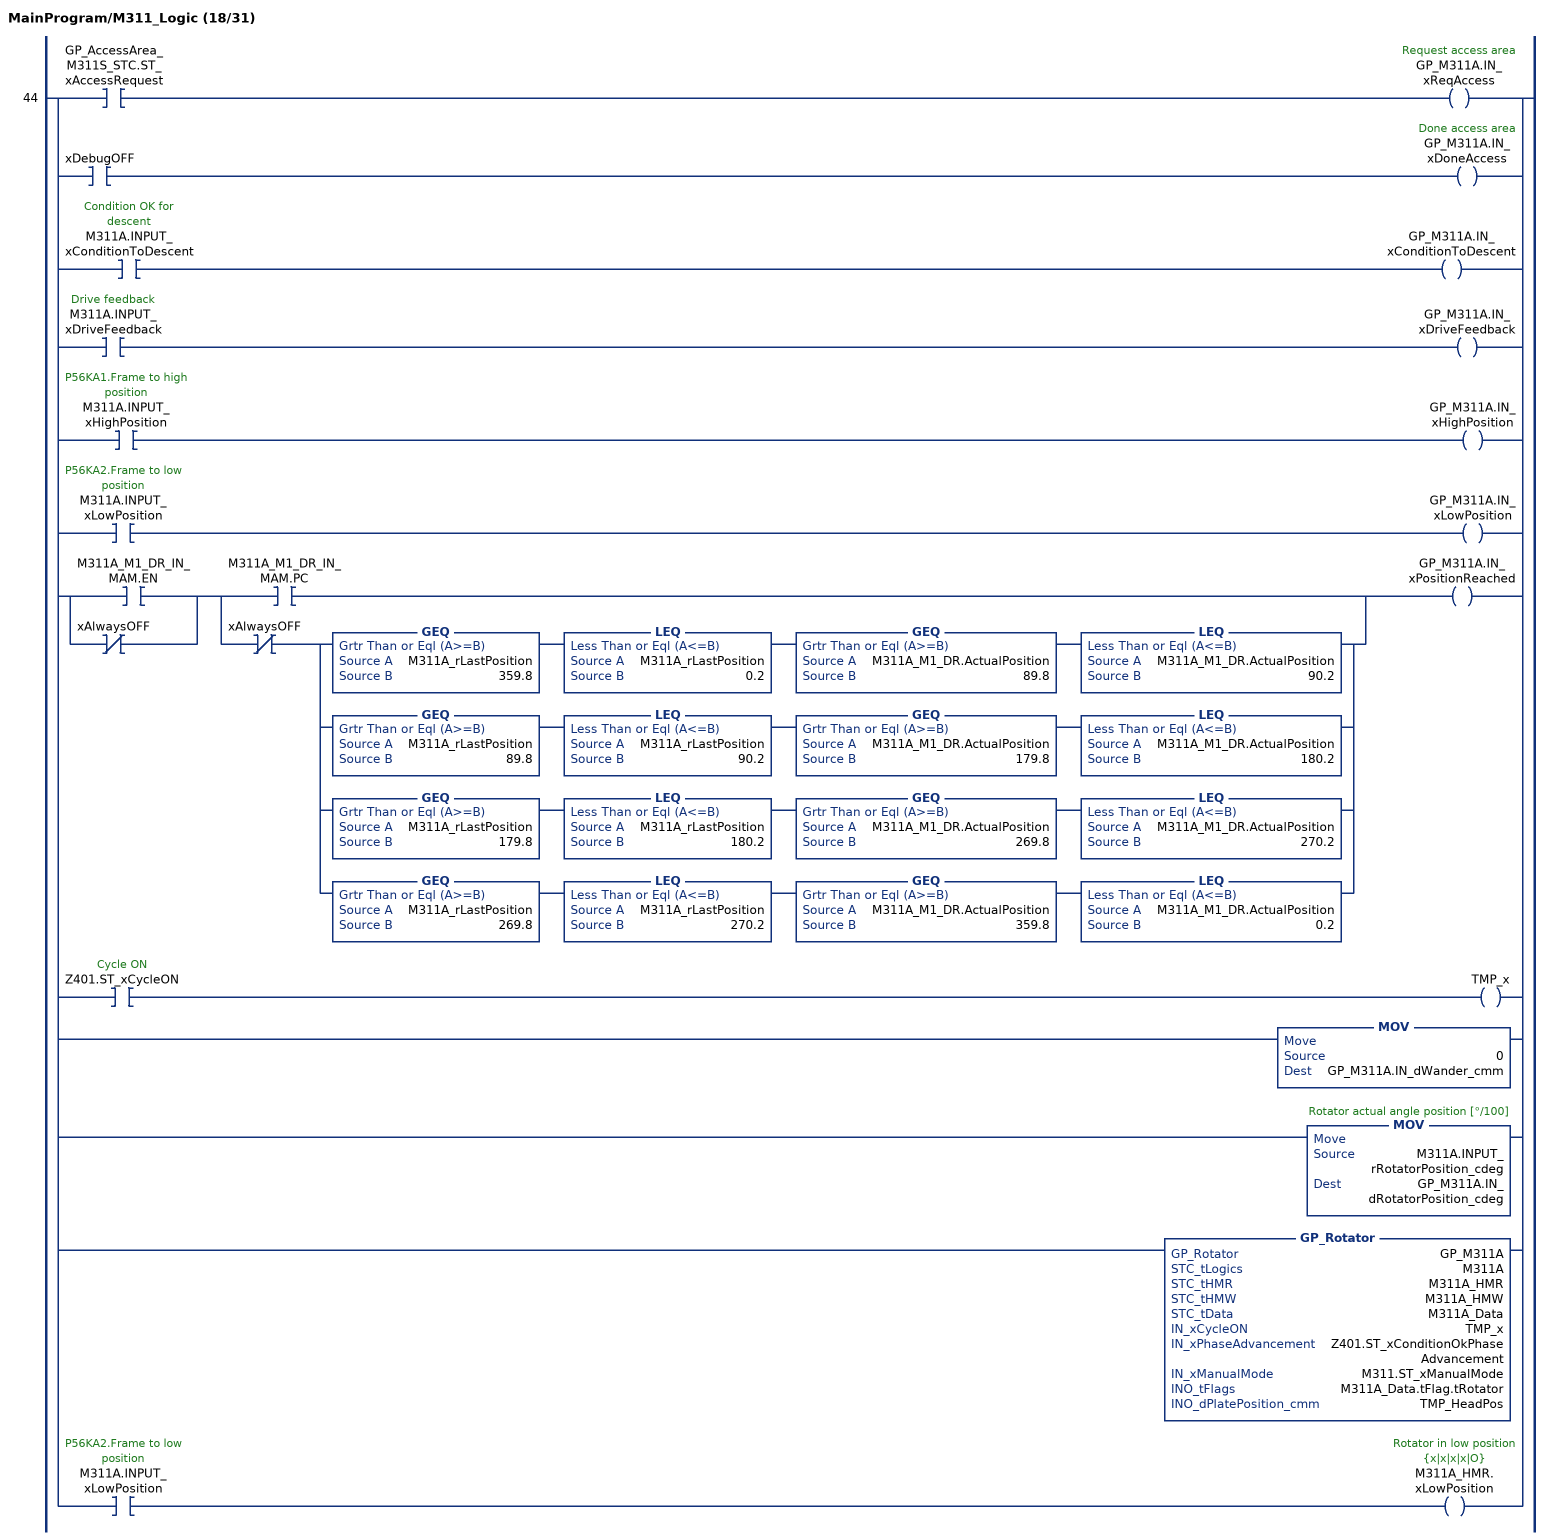
   44: [XIC(GP_AccessArea_M311S_STC.ST_xAccessRequest) OTE(GP_M311A.IN_xReqAccess) ,XIC(xDebugOFF) OTE(GP_M311A.IN_xDoneAccess) ,XIC(M311A.INPUT_xConditionToDescent) OTE(GP_M311A.IN_xConditionToDescent) ,XIC(M311A.INPUT_xDriveFeedback) OTE(GP_M311A.IN_xDriveFeedback) ,XIC(M311A.INPUT_xHighPosition) OTE(GP_M311A.IN_xHighPosition) ,XIC(M311A.INPUT_xLowPosition) OTE(GP_M311A.IN_xLowPosition) ,[XIC(M311A_M1_DR_IN_MAM.EN) ,XIO(xAlwaysOFF) ] [XIC(M311A_M1_DR_IN_MAM.PC) ,XIO(xAlwaysOFF) [GEQ(M311A_rLastPosition,359.8) LEQ(M311A_rLastPosition,0.2) GEQ(M311A_M1_DR.ActualPosition,89.8) LEQ(M311A_M1_DR.ActualPosition,90.2) ,GEQ(M311A_rLastPosition,89.8) LEQ(M311A_rLastPosition,90.2) GEQ(M311A_M1_DR.ActualPosition,179.8) LEQ(M311A_M1_DR.ActualPosition,180.2) ,GEQ(M311A_rLastPosition,179.8) LEQ(M311A_rLastPosition,180.2) GEQ(M311A_M1_DR.ActualPosition,269.8) LEQ(M311A_M1_DR.ActualPosition,270.2) ,GEQ(M311A_rLastPosition,269.8) LEQ(M311A_rLastPosition,270.2) GEQ(M311A_M1_DR.ActualPosition,359.8) LEQ(M311A_M1_DR.ActualPosition,0.2) ] ] OTE(GP_M311A.IN_xPositionReached) ,XIC(Z401.ST_xCycleON) OTE(TMP_x) ,MOV(0,GP_M311A.IN_dWander_cmm) ,MOV(M311A.INPUT_rRotatorPosition_cdeg,GP_M311A.IN_dRotatorPosition_cdeg) ,GP_Rotator(GP_M311A,M311A,M311A_HMR,M311A_HMW,M311A_Data,TMP_x,Z401.ST_xConditionOkPhaseAdvancement,M311.ST_xManualMode,M311A_Data.tFlag.tRotator,TMP_HeadPos) ,XIC(M311A.INPUT_xLowPosition) OTE(M311A_HMR.xLowPosition) ];
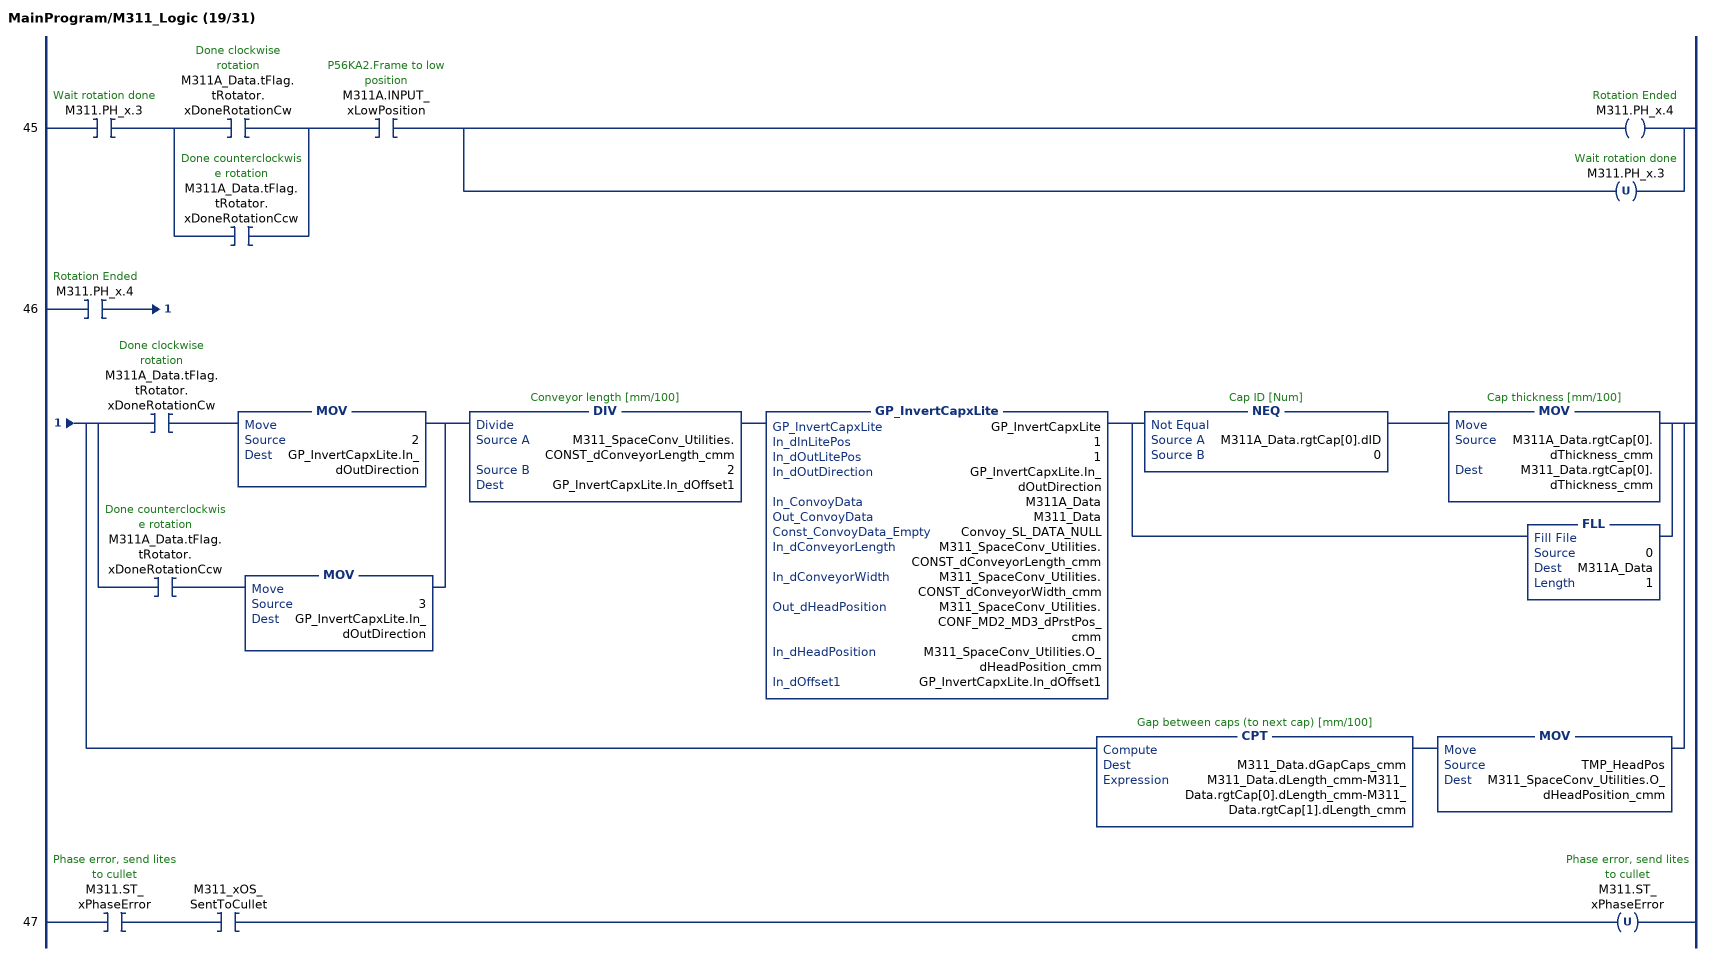
   45: XIC(M311.PH_x.3)[XIC(M311A_Data.tFlag.tRotator.xDoneRotationCw) ,XIC(M311A_Data.tFlag.tRotator.xDoneRotationCcw) ]XIC(M311A.INPUT_xLowPosition)[OTE(M311.PH_x.4) ,OTU(M311.PH_x.3) ];
   46: XIC(M311.PH_x.4)[[XIC(M311A_Data.tFlag.tRotator.xDoneRotationCw) MOV(2,GP_InvertCapxLite.In_dOutDirection) ,XIC(M311A_Data.tFlag.tRotator.xDoneRotationCcw) MOV(3,GP_InvertCapxLite.In_dOutDirection) ] DIV(M311_SpaceConv_Utilities.CONST_dConveyorLength_cmm,2,GP_InvertCapxLite.In_dOffset1) GP_InvertCapxLite(GP_InvertCapxLite,1,1,GP_InvertCapxLite.In_dOutDirection,M311A_Data,M311_Data,Convoy_SL_DATA_NULL,M311_SpaceConv_Utilities.CONST_dConveyorLength_cmm,M311_SpaceConv_Utilities.CONST_dConveyorWidth_cmm,M311_SpaceConv_Utilities.CONF_MD2_MD3_dPrstPos_cmm,M311_SpaceConv_Utilities.O_dHeadPosition_cmm,GP_InvertCapxLite.In_dOffset1) [NEQ(M311A_Data.rgtCap[0].dID,0) MOV(M311A_Data.rgtCap[0].dThickness_cmm,M311_Data.rgtCap[0].dThickness_cmm) ,FLL(0,M311A_Data,1) ] ,CPT(M311_Data.dGapCaps_cmm,M311_Data.dLength_cmm-M311_Data.rgtCap[0].dLength_cmm-M311_Data.rgtCap[1].dLength_cmm) MOV(TMP_HeadPos,M311_SpaceConv_Utilities.O_dHeadPosition_cmm) ];
   47: XIC(M311.ST_xPhaseError)XIC(M311_xOS_SentToCullet)OTU(M311.ST_xPhaseError);
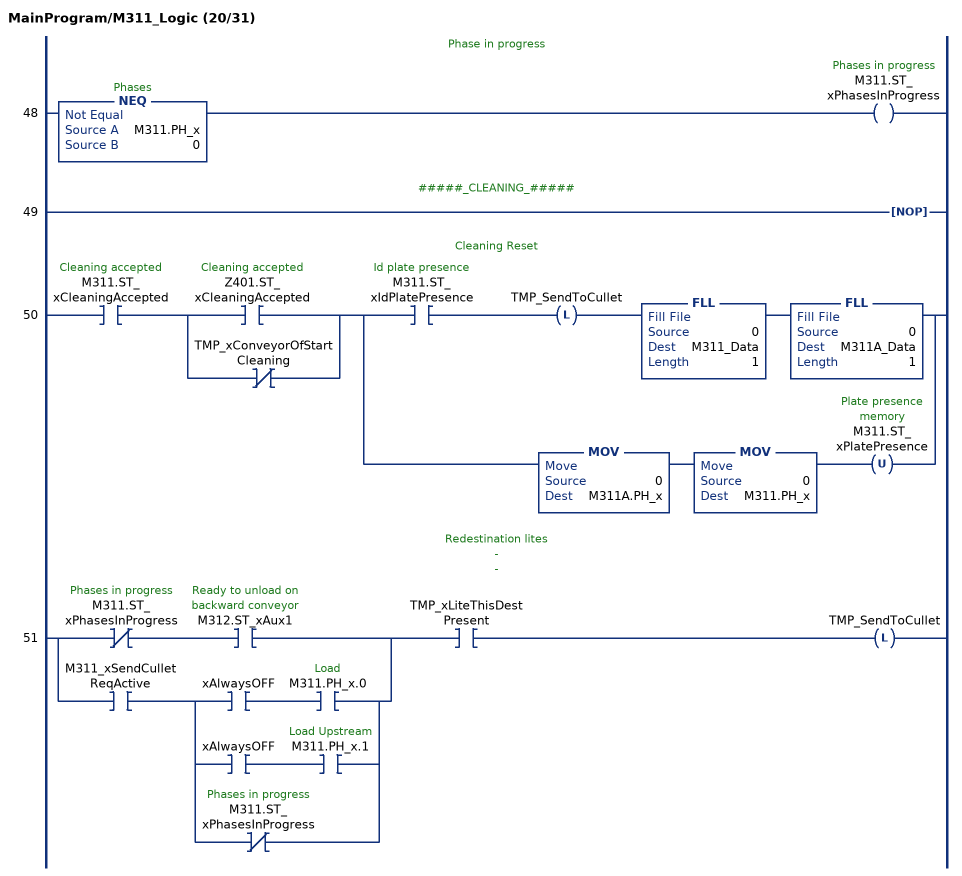
   // Phase in progress
   48: NEQ(M311.PH_x,0)OTE(M311.ST_xPhasesInProgress);
   // #####_CLEANING_#####
   49: NOP();
   // Cleaning Reset
   50: XIC(M311.ST_xCleaningAccepted)[XIC(Z401.ST_xCleaningAccepted) ,XIO(TMP_xConveyorOfStartCleaning) ][XIC(M311.ST_xIdPlatePresence) OTL(TMP_SendToCullet) FLL(0,M311_Data,1) FLL(0,M311A_Data,1) ,MOV(0,M311A.PH_x) MOV(0,M311.PH_x) OTU(M311.ST_xPlatePresence) ];
   // Redestination lites
   // -
   // -
   51: [XIO(M311.ST_xPhasesInProgress) XIC(M312.ST_xAux1) ,XIC(M311_xSendCulletReqActive) [XIC(xAlwaysOFF) XIC(M311.PH_x.0) ,XIC(xAlwaysOFF) XIC(M311.PH_x.1) ,XIO(M311.ST_xPhasesInProgress) ] ]XIC(TMP_xLiteThisDestPresent)OTL(TMP_SendToCullet);
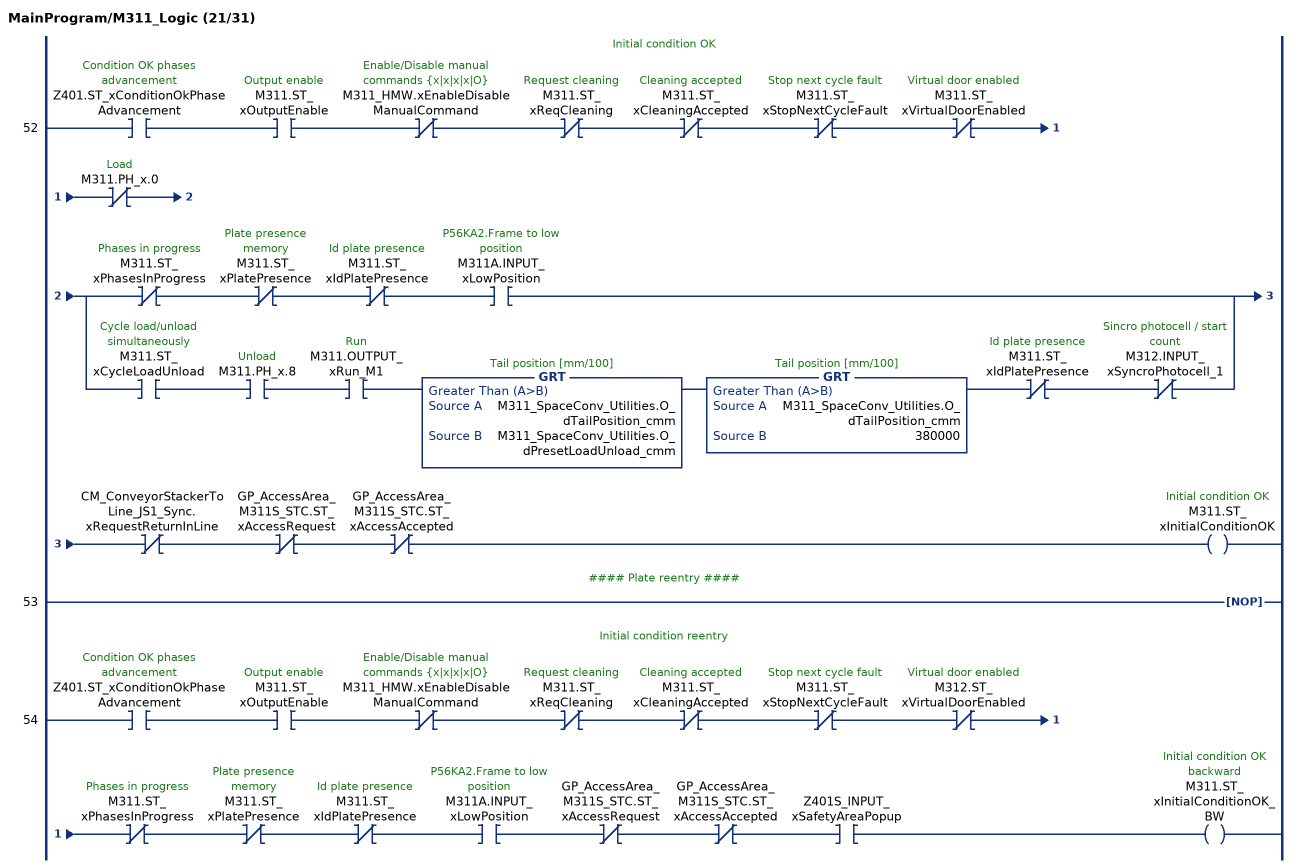
   // Initial condition OK
   52: XIC(Z401.ST_xConditionOkPhaseAdvancement)XIC(M311.ST_xOutputEnable)XIO(M311_HMW.xEnableDisableManualCommand)XIO(M311.ST_xReqCleaning)XIO(M311.ST_xCleaningAccepted)XIO(M311.ST_xStopNextCycleFault)XIO(M311.ST_xVirtualDoorEnabled)XIO(M311.PH_x.0)[XIO(M311.ST_xPhasesInProgress) XIO(M311.ST_xPlatePresence) XIO(M311.ST_xIdPlatePresence) XIC(M311A.INPUT_xLowPosition) ,XIC(M311.ST_xCycleLoadUnload) XIC(M311.PH_x.8) XIC(M311.OUTPUT_xRun_M1) GRT(M311_SpaceConv_Utilities.O_dTailPosition_cmm,M311_SpaceConv_Utilities.O_dPresetLoadUnload_cmm) GRT(M311_SpaceConv_Utilities.O_dTailPosition_cmm,380000) XIO(M311.ST_xIdPlatePresence) XIO(M312.INPUT_xSyncroPhotocell_1) ]XIO(CM_ConveyorStackerToLine_JS1_Sync.xRequestReturnInLine)XIO(GP_AccessArea_M311S_STC.ST_xAccessRequest)XIO(GP_AccessArea_M311S_STC.ST_xAccessAccepted)OTE(M311.ST_xInitialConditionOK);
   // #### Plate reentry ####
   53: NOP();
   // Initial condition reentry
   54: XIC(Z401.ST_xConditionOkPhaseAdvancement)XIC(M311.ST_xOutputEnable)XIO(M311_HMW.xEnableDisableManualCommand)XIO(M311.ST_xReqCleaning)XIO(M311.ST_xCleaningAccepted)XIO(M311.ST_xStopNextCycleFault)XIO(M312.ST_xVirtualDoorEnabled)XIO(M311.ST_xPhasesInProgress)XIO(M311.ST_xPlatePresence)XIO(M311.ST_xIdPlatePresence)XIC(M311A.INPUT_xLowPosition)XIO(GP_AccessArea_M311S_STC.ST_xAccessRequest)XIO(GP_AccessArea_M311S_STC.ST_xAccessAccepted)XIC(Z401S_INPUT_xSafetyAreaPopup)OTE(M311.ST_xInitialConditionOK_BW);
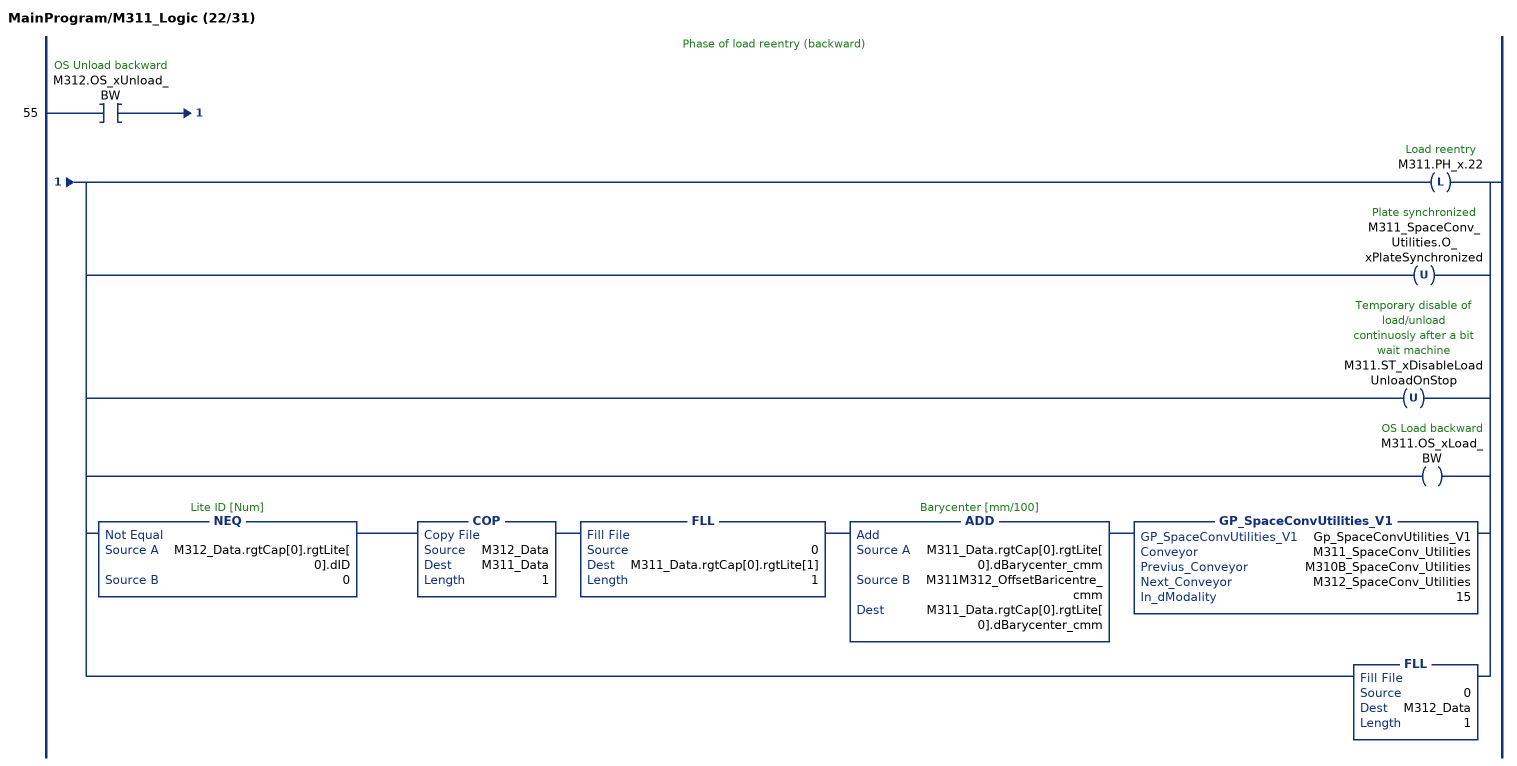
   // Phase of load reentry (backward)
   55: XIC(M312.OS_xUnload_BW)[OTL(M311.PH_x.22) ,OTU(M311_SpaceConv_Utilities.O_xPlateSynchronized) ,OTU(M311.ST_xDisableLoadUnloadOnStop) ,OTE(M311.OS_xLoad_BW) ,NEQ(M312_Data.rgtCap[0].rgtLite[0].dID,0) COP(M312_Data,M311_Data,1) FLL(0,M311_Data.rgtCap[0].rgtLite[1],1) ADD(M311_Data.rgtCap[0].rgtLite[0].dBarycenter_cmm,M311M312_OffsetBaricentre_cmm,M311_Data.rgtCap[0].rgtLite[0].dBarycenter_cmm) GP_SpaceConvUtilities_V1(Gp_SpaceConvUtilities_V1,M311_SpaceConv_Utilities,M310B_SpaceConv_Utilities,M312_SpaceConv_Utilities,15) ,FLL(0,M312_Data,1) ];
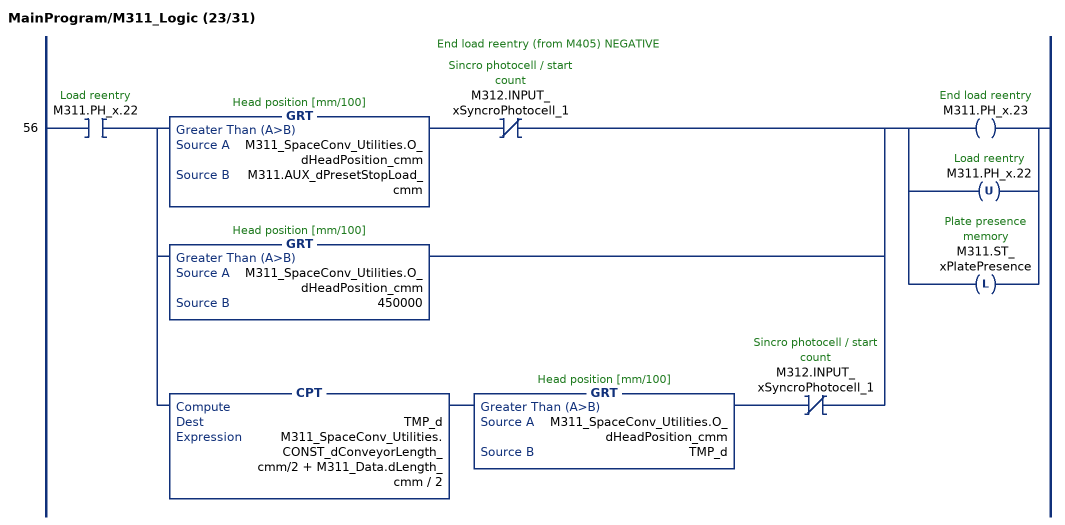
   // End load reentry (from M405) NEGATIVE
   56: XIC(M311.PH_x.22)[[GRT(M311_SpaceConv_Utilities.O_dHeadPosition_cmm,M311.AUX_dPresetStopLoad_cmm) XIO(M312.INPUT_xSyncroPhotocell_1) ,GRT(M311_SpaceConv_Utilities.O_dHeadPosition_cmm,450000) ] ,CPT(TMP_d,M311_SpaceConv_Utilities.CONST_dConveyorLength_cmm/2 + M311_Data.dLength_cmm / 2) GRT(M311_SpaceConv_Utilities.O_dHeadPosition_cmm,TMP_d) XIO(M312.INPUT_xSyncroPhotocell_1) ][OTE(M311.PH_x.23) ,OTU(M311.PH_x.22) ,OTL(M311.ST_xPlatePresence) ];
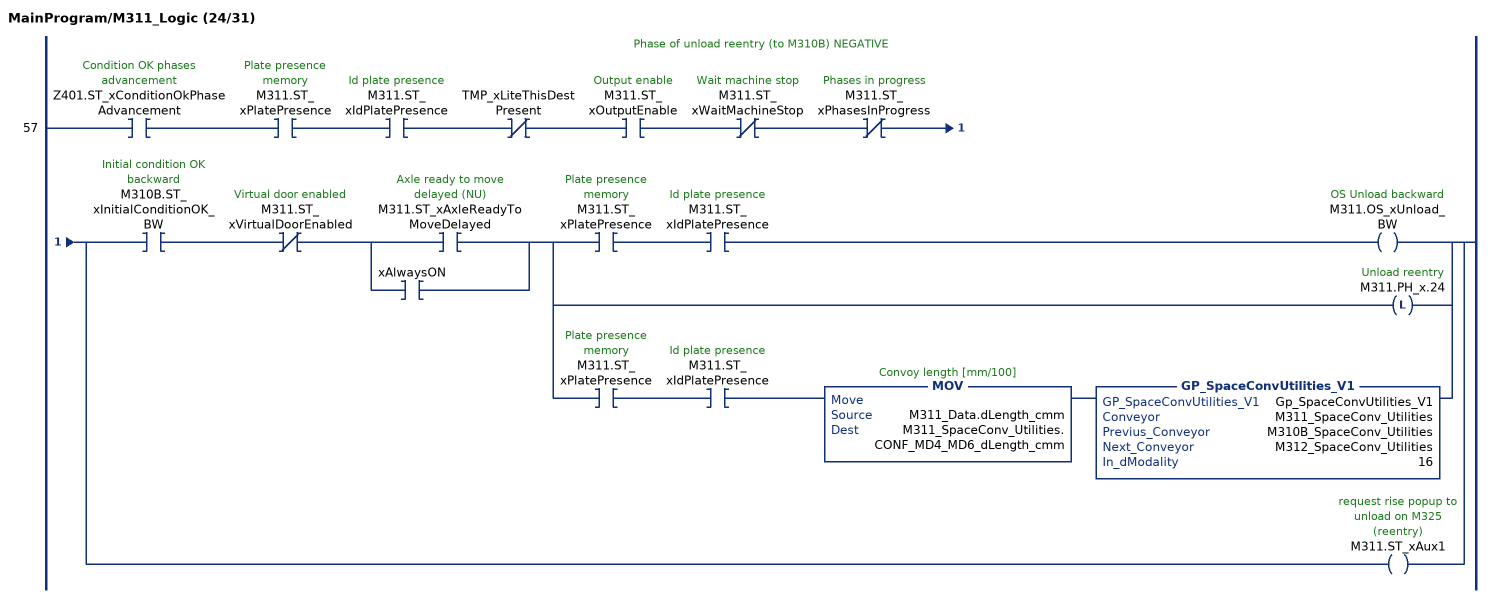
   // Phase of unload reentry (to M310B) NEGATIVE
   57: XIC(Z401.ST_xConditionOkPhaseAdvancement)XIC(M311.ST_xPlatePresence)XIC(M311.ST_xIdPlatePresence)XIO(TMP_xLiteThisDestPresent)XIC(M311.ST_xOutputEnable)XIO(M311.ST_xWaitMachineStop)XIO(M311.ST_xPhasesInProgress)[XIC(M310B.ST_xInitialConditionOK_BW) XIO(M311.ST_xVirtualDoorEnabled) [XIC(M311.ST_xAxleReadyToMoveDelayed) ,XIC(xAlwaysON) ] [XIC(M311.ST_xPlatePresence) XIC(M311.ST_xIdPlatePresence) OTE(M311.OS_xUnload_BW) ,OTL(M311.PH_x.24) ,XIC(M311.ST_xPlatePresence) XIC(M311.ST_xIdPlatePresence) MOV(M311_Data.dLength_cmm,M311_SpaceConv_Utilities.CONF_MD4_MD6_dLength_cmm) GP_SpaceConvUtilities_V1(Gp_SpaceConvUtilities_V1,M311_SpaceConv_Utilities,M310B_SpaceConv_Utilities,M312_SpaceConv_Utilities,16) ] ,OTE(M311.ST_xAux1) ];
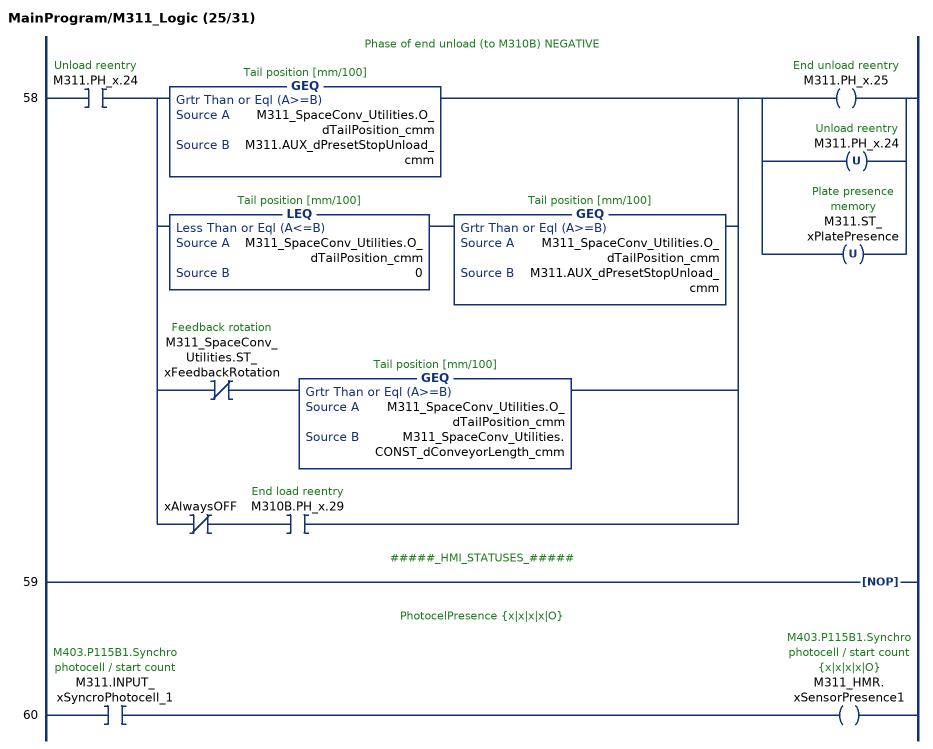
   // Phase of end unload (to M310B) NEGATIVE
   58: XIC(M311.PH_x.24)[[GEQ(M311_SpaceConv_Utilities.O_dTailPosition_cmm,M311.AUX_dPresetStopUnload_cmm) ,LEQ(M311_SpaceConv_Utilities.O_dTailPosition_cmm,0) GEQ(M311_SpaceConv_Utilities.O_dTailPosition_cmm,M311.AUX_dPresetStopUnload_cmm) ] ,XIO(M311_SpaceConv_Utilities.ST_xFeedbackRotation) GEQ(M311_SpaceConv_Utilities.O_dTailPosition_cmm,M311_SpaceConv_Utilities.CONST_dConveyorLength_cmm) ,XIO(xAlwaysOFF) XIC(M310B.PH_x.29) ][OTE(M311.PH_x.25) ,OTU(M311.PH_x.24) ,OTU(M311.ST_xPlatePresence) ];
   // #####_HMI_STATUSES_#####
   59: NOP();
   // PhotocelPresence {x|x|x|x|O}
   60: XIC(M311.INPUT_xSyncroPhotocell_1)OTE(M311_HMR.xSensorPresence1);
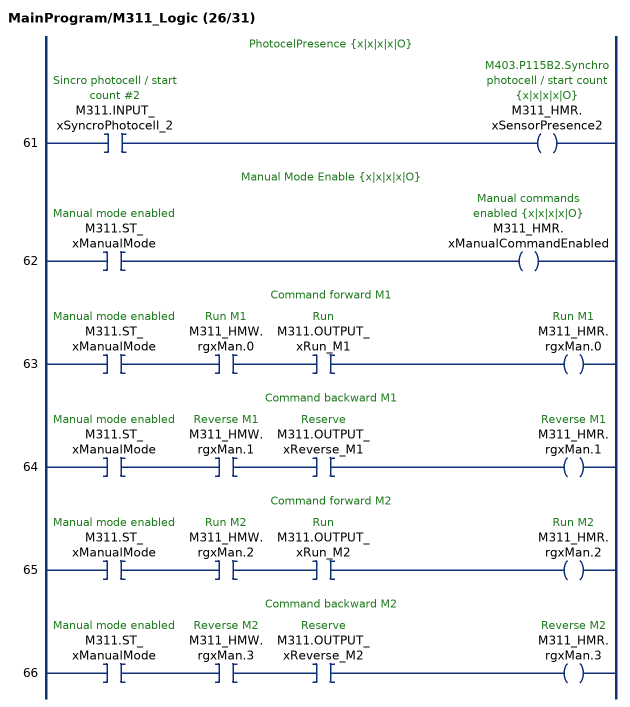
   // PhotocelPresence {x|x|x|x|O}
   61: XIC(M311.INPUT_xSyncroPhotocell_2)OTE(M311_HMR.xSensorPresence2);
   // Manual Mode Enable {x|x|x|x|O}
   62: XIC(M311.ST_xManualMode)OTE(M311_HMR.xManualCommandEnabled);
   // Command forward M1
   63: XIC(M311.ST_xManualMode)XIC(M311_HMW.rgxMan.0)XIC(M311.OUTPUT_xRun_M1)OTE(M311_HMR.rgxMan.0);
   // Command backward M1
   64: XIC(M311.ST_xManualMode)XIC(M311_HMW.rgxMan.1)XIC(M311.OUTPUT_xReverse_M1)OTE(M311_HMR.rgxMan.1);
   // Command forward M2
   65: XIC(M311.ST_xManualMode)XIC(M311_HMW.rgxMan.2)XIC(M311.OUTPUT_xRun_M2)OTE(M311_HMR.rgxMan.2);
   // Command backward M2
   66: XIC(M311.ST_xManualMode)XIC(M311_HMW.rgxMan.3)XIC(M311.OUTPUT_xReverse_M2)OTE(M311_HMR.rgxMan.3);
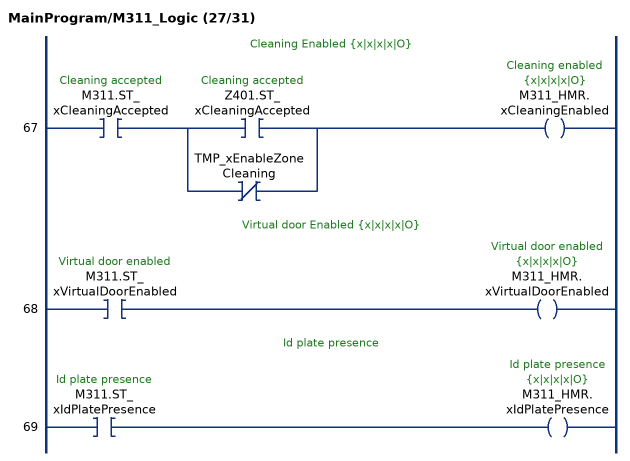
   // Cleaning Enabled {x|x|x|x|O}
   67: XIC(M311.ST_xCleaningAccepted)[XIC(Z401.ST_xCleaningAccepted) ,XIO(TMP_xEnableZoneCleaning) ]OTE(M311_HMR.xCleaningEnabled);
   // Virtual door Enabled {x|x|x|x|O}
   68: XIC(M311.ST_xVirtualDoorEnabled)OTE(M311_HMR.xVirtualDoorEnabled);
   // Id plate presence
   69: XIC(M311.ST_xIdPlatePresence)OTE(M311_HMR.xIdPlatePresence);
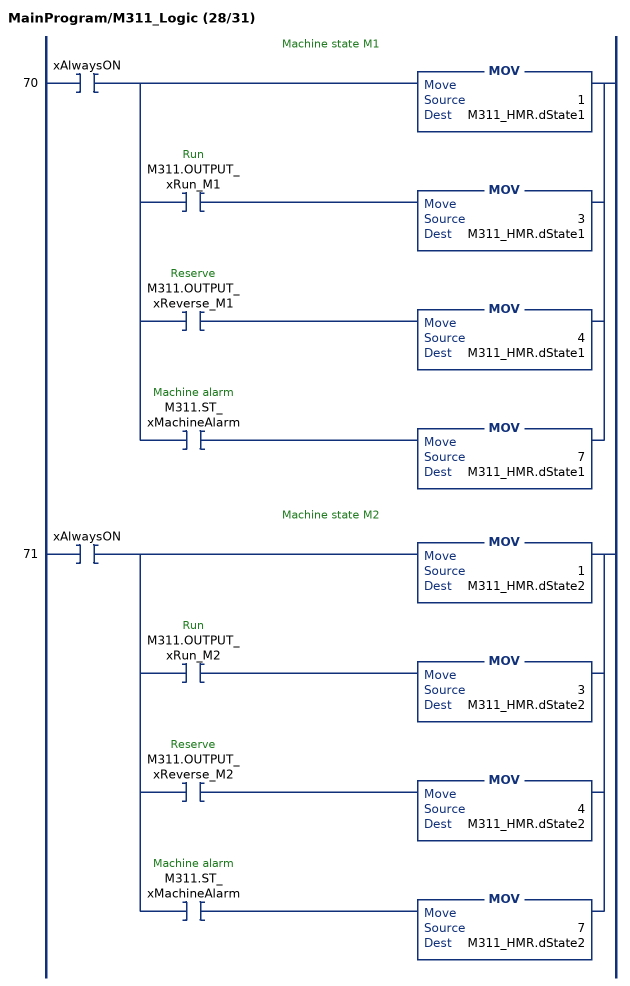
   // Machine state M1
   70: XIC(xAlwaysON)[MOV(1,M311_HMR.dState1) ,XIC(M311.OUTPUT_xRun_M1) MOV(3,M311_HMR.dState1) ,XIC(M311.OUTPUT_xReverse_M1) MOV(4,M311_HMR.dState1) ,XIC(M311.ST_xMachineAlarm) MOV(7,M311_HMR.dState1) ];
   // Machine state M2
   71: XIC(xAlwaysON)[MOV(1,M311_HMR.dState2) ,XIC(M311.OUTPUT_xRun_M2) MOV(3,M311_HMR.dState2) ,XIC(M311.OUTPUT_xReverse_M2) MOV(4,M311_HMR.dState2) ,XIC(M311.ST_xMachineAlarm) MOV(7,M311_HMR.dState2) ];
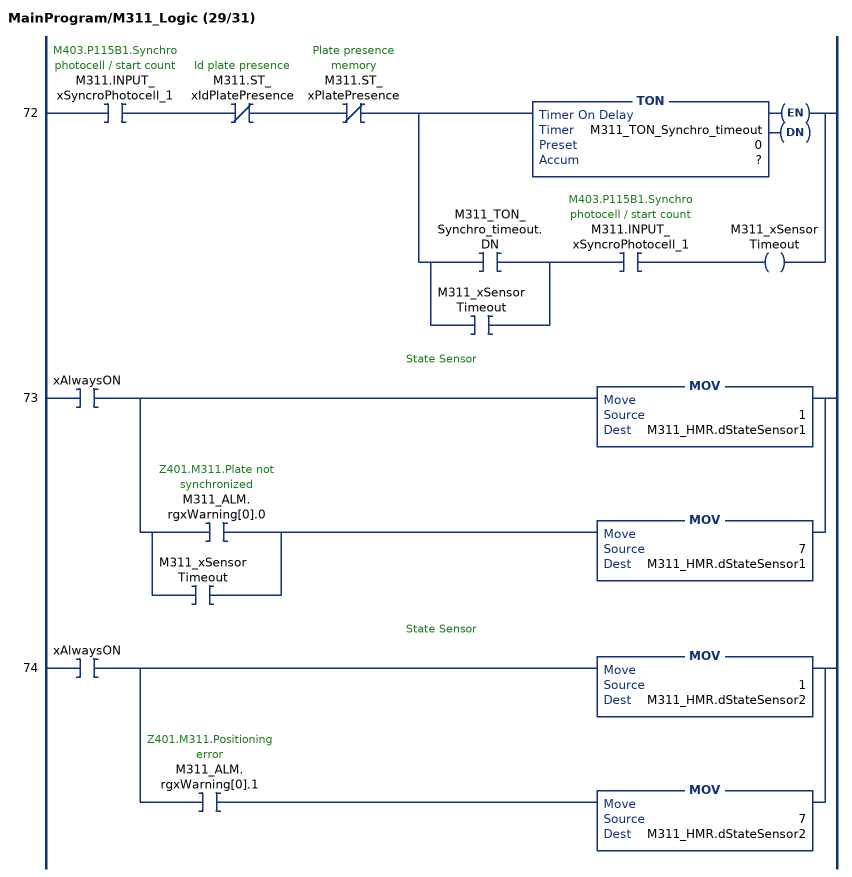
   72: XIC(M311.INPUT_xSyncroPhotocell_1)XIO(M311.ST_xIdPlatePresence)XIO(M311.ST_xPlatePresence)[TON(M311_TON_Synchro_timeout,?,?) ,[XIC(M311_TON_Synchro_timeout.DN) ,XIC(M311_xSensorTimeout) ] XIC(M311.INPUT_xSyncroPhotocell_1) OTE(M311_xSensorTimeout) ];
   // State Sensor
   73: XIC(xAlwaysON)[MOV(1,M311_HMR.dStateSensor1) ,[XIC(M311_ALM.rgxWarning[0].0) ,XIC(M311_xSensorTimeout) ] MOV(7,M311_HMR.dStateSensor1) ];
   // State Sensor
   74: XIC(xAlwaysON)[MOV(1,M311_HMR.dStateSensor2) ,XIC(M311_ALM.rgxWarning[0].1) MOV(7,M311_HMR.dStateSensor2) ];
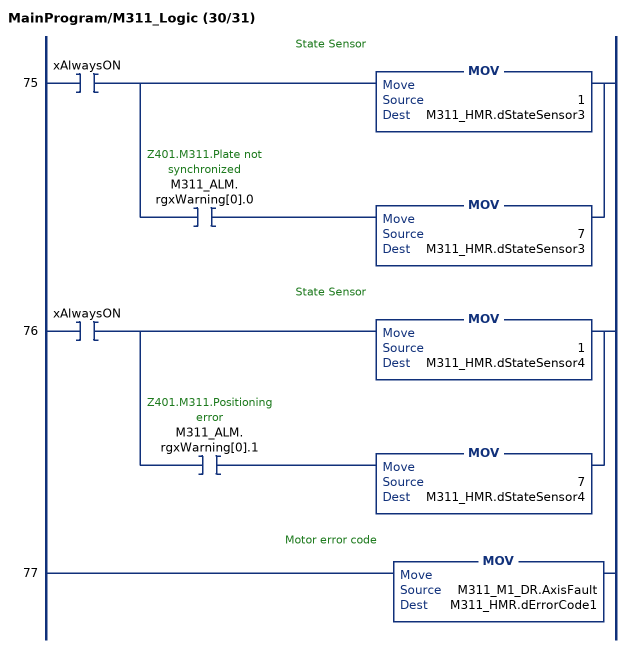
   // State Sensor
   75: XIC(xAlwaysON)[MOV(1,M311_HMR.dStateSensor3) ,XIC(M311_ALM.rgxWarning[0].0) MOV(7,M311_HMR.dStateSensor3) ];
   // State Sensor
   76: XIC(xAlwaysON)[MOV(1,M311_HMR.dStateSensor4) ,XIC(M311_ALM.rgxWarning[0].1) MOV(7,M311_HMR.dStateSensor4) ];
   // Motor error code
   77: MOV(M311_M1_DR.AxisFault,M311_HMR.dErrorCode1);
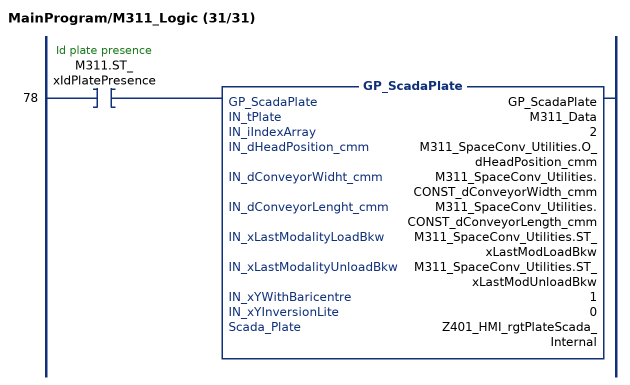
   78: XIC(M311.ST_xIdPlatePresence)GP_ScadaPlate(GP_ScadaPlate,M311_Data,2,M311_SpaceConv_Utilities.O_dHeadPosition_cmm,M311_SpaceConv_Utilities.CONST_dConveyorWidth_cmm,M311_SpaceConv_Utilities.CONST_dConveyorLength_cmm,M311_SpaceConv_Utilities.ST_xLastModLoadBkw,M311_SpaceConv_Utilities.ST_xLastModUnloadBkw,1,0,Z401_HMI_rgtPlateScada_Internal);
END_ROUTINE
